(* Logix 5000 project; controller FV vendor 1 type 14 code 217 rev 31.11; software revision 31.00; part 54 of 63 *)
(* tags used below, declared in another part *)
   Alarm_Reset : BOOL;
   CWD : CHECKWORD_FLAGS;
   Default_Check_Time : DINT;
   Dummy : BOOL;
   FV_AV1 : PlantItem;   // AV1
   FV_AV1_ALARM : ALARM_DIGITAL;
   FV_AV1_C : ALIAS FOR Remote_IO:6:I.Data.4;   // YSV 1 outlet valve closed f/b
   FV_AV1_DR : ALIAS FOR Remote_IO:5:O.Data.0;   // YSV 1 outlet valve
   FV_AV1_O : ALIAS FOR Remote_IO:6:I.Data.0;   // YSV 1 outlet valve open f/b
   FV_AV1A : PlantItem;   // AV1A
   FV_AV1A_ALARM : ALARM_DIGITAL;
   FV_AV1A_C : ALIAS FOR Remote_IO:6:I.Data.10;   // AV1A seat clean valve closed f/b
   FV_AV1A_DR : ALIAS FOR Remote_IO:5:O.Data.4;   // AV1 seat clean valve
   FV_AV1A_O : ALIAS FOR Remote_IO:6:I.Data.8;   // AV1A seat clean valve open f/b
   FV_AV2 : PlantItem;   // AV2
   FV_AV2_ALARM : ALARM_DIGITAL;
   FV_AV2_C : ALIAS FOR Remote_IO:6:I.Data.5;   // Water flush valve closed f/b
   FV_AV2_DR : ALIAS FOR Remote_IO:5:O.Data.1;   // Water flush valve
   FV_AV2_O : ALIAS FOR Remote_IO:6:I.Data.1;   // Water flush valve open f/b
   FV_AV3 : PlantItem;   // AV3
   FV_AV3_ALARM : ALARM_DIGITAL;
   FV_AV3_C : ALIAS FOR Remote_IO:6:I.Data.6;   // CIP delivery valve closed f/b
   FV_AV3_DR : ALIAS FOR Remote_IO:5:O.Data.2;   // CIP delivery valve
   FV_AV3_O : ALIAS FOR Remote_IO:6:I.Data.2;   // CIP delivery valve open f/b
   FV_AV4 : PlantItem;   // AV4
   FV_AV4_ALARM : ALARM_DIGITAL;
   FV_AV4_C : ALIAS FOR Remote_IO:6:I.Data.7;   // Centrifuge main closed f/b
   FV_AV4_DR : ALIAS FOR Remote_IO:5:O.Data.3;   // Centrifuge main valve
   FV_AV4_O : ALIAS FOR Remote_IO:6:I.Data.3;   // Centrifuge main valve f/b
   FV_AV4A : PlantItem;   // AV4A
   FV_AV4A_ALARM : ALARM_DIGITAL;
   FV_AV4A_C : ALIAS FOR Remote_IO:6:I.Data.11;   // AV4A seat clean valve closed f/b
   FV_AV4A_DR : ALIAS FOR Remote_IO:5:O.Data.5;   // AV4 seat clean valve
   FV_AV4A_O : ALIAS FOR Remote_IO:6:I.Data.9;   // AV4A seat clean valve closed f/b
   FV_AV5 : PlantItem;   // AV5
   FV_AV5_ALARM : ALARM_DIGITAL;
   FV_AV5_C : ALIAS FOR Remote_IO:7:I.Data.9;
   FV_AV5_DR : ALIAS FOR Remote_IO:9:O.Data.12;
   FV_AV5_O : ALIAS FOR Remote_IO:7:I.Data.8;
   FV_B17 : INT[255];   // VES_ACTIVE Vessel active flags
   fv_bit_data_file_address : INT;
   fv_bit_file_bit_offset : INT;
   fv_bit_file_word_offset : INT;
   fv_bit_offset : INT;
   fv_bit_value_to_set : INT;
   FV_data_file_address : INT;
   FV_N110 : INT[255];   // FV DATA 0 CURRENT FV DATA
   FV_N111 : INT[50];   // FV1, CURRENT FV DATA
   FV_N112 : INT[50];   // FV2, CURRENT FV DATA
   FV_N113 : INT[50];   // FV3, CURRENT FV DATA
   FV_N114 : INT[50];   // FV4, CURRENT FV DATA
   FV_N115 : INT[50];   // FV5, CURRENT FV DATA
   FV_N116 : INT[50];   // FV6, CURRENT FV DATA
   FV_N117 : INT[50];   // FV7, CURRENT FV DATA
   FV_N118 : INT[50];   // FV8, CURRENT FV DATA
   FV_N119 : INT[50];   // FV9, CURRENT FV DATA
   FV_N120 : INT[50];   // FV10, CURRENT FV DATA
   FV_N121 : INT[50];   // FV11, CURRENT FV DATA
   FV_N122 : INT[50];   // FV12, CURRENT FV DATA
   FV_N123 : INT[50];   // FV13, CURRENT FV DATA
   FV_N124 : INT[50];   // FV14, CURRENT FV DATA
   FV_N125 : INT[50];   // FV15, CURRENT FV DATA
   FV_N126 : INT[50];   // FV16, CURRENT FV DATA
   FV_N127 : INT[50];   // FV17, CURRENT FV DATA
   FV_N128 : INT[50];   // FV18, CURRENT FV DATA
   FV_N129 : INT[50];   // FV19, CURRENT FV DATA
   FV_N130 : INT[50];   // FV20, CURRENT FV DATA
   FV_N131 : INT[50];   // FV21, CURRENT FV DATA
   FV_N132 : INT[50];   // FV22, CURRENT FV DATA
   FV_N133 : INT[50];   // FV23, CURRENT FV DATA
   FV_N134 : INT[50];   // FV24, CURRENT FV DATA
   FV_N135 : INT[50];   // FV25, CURRENT FV DATA
   FV_N136 : INT[50];   // YSV1, CURRENT FV DATA
   FV_N137 : INT[50];   // YSV2, CURRENT FV DATA
   FV_N138 : INT[50];   // YSV3, CURRENT FV DATA
   FV_N139 : INT[255];   // YST1
   FV_N140 : INT[255];   // YST2
   FV_N141 : INT[255];   // YSV1 DATA
   FV_N142 : INT[255];   // YSV2 DATA
   FV_N143 : INT[255];   // YSV3 DATA
   FV_N144 : INT[255];   // YST1 DATA
   FV_N145 : INT[255];   // YST2 DATA
   FV_N146 : INT[50];   // FV26, CURRENT FV DATA
   FV_N147 : INT[50];   // FV27, CURRENT FV DATA
   FV_N148 : INT[50];   // FV28, CURRENT FV DATA
   FV_N149 : INT[50];   // FV29, CURRENT FV DATA
   FV_N150 : INT[50];   // FV30, CURRENT FV DATA
   FV_N151 : INT[50];   // FV31, CURRENT FV DATA
   FV_R2V1 : PlantItem;   // R2V1
   FV_R2V1_ALARM : ALARM_DIGITAL;
   FV_R2V1_C : ALIAS FOR Remote_IO:7:I.Data.6;
   FV_R2V1_DR : ALIAS FOR Remote_IO:5:O.Data.10;
   FV_R2V1_O : ALIAS FOR Remote_IO:7:I.Data.2;
   FV_R2V2 : PlantItem;   // R2V2
   FV_R2V2_ALARM : ALARM_DIGITAL;
   FV_R2V2_C : ALIAS FOR Remote_IO:7:I.Data.7;
   FV_R2V2_DR : ALIAS FOR Remote_IO:5:O.Data.11;
   FV_R2V2_O : ALIAS FOR Remote_IO:7:I.Data.3;
   FV_value_to_set : INT;
   FV_word_offset : INT;
   FV_WYTR1 : PlantItem;   // WYTR1
   FV_WYTR1_ALARM : ALARM_DIGITAL;
   FV_WYTR1_C : ALIAS FOR Remote_IO:7:I.Data.4;
   FV_WYTR1_DR : ALIAS FOR Remote_IO:5:O.Data.8;
   FV_WYTR1_O : ALIAS FOR Remote_IO:7:I.Data.0;
   FV_WYTR2 : PlantItem;   // WYTR2
   FV_WYTR2_ALARM : ALARM_DIGITAL;
   FV_WYTR2_C : ALIAS FOR Remote_IO:7:I.Data.5;
   FV_WYTR2_DR : ALIAS FOR Remote_IO:5:O.Data.9;
   FV_WYTR2_O : ALIAS FOR Remote_IO:7:I.Data.1;
   Item_Faults_Are_Latched : BOOL;
   Item_Simulation_Flag : BOOL;
   One_Second_One_Scan : ALIAS FOR One_Second_1_scan;
   Scada_Valve_Fault_No : DINT;
   YP_AV2 : PlantItem;   // AV2
   YP_AV2_ALARM : ALARM_DIGITAL;
   YP_AV2_DR : ALIAS FOR RIO_Rack_3:3:O.Data.5;
   YP_AV2_O : ALIAS FOR RIO_Rack_3:1:I.Data.2;
(* FV_Common, continued *)

ROUTINE FV_Set_FV_Datafile_Value   (* ladder *)
   // Routine to Set the value of something within the FV Data Files, Used to replace indirection originally used
   0: SBR(FV_value_to_set,FV_data_file_address,FV_word_offset)OTE(Dummy);
   1: EQU(FV_data_file_address,110)MOV(FV_value_to_set,FV_N110[FV_word_offset]);
   2: EQU(FV_data_file_address,111)MOV(FV_value_to_set,FV_N111[FV_word_offset]);
   3: EQU(FV_data_file_address,112)MOV(FV_value_to_set,FV_N112[FV_word_offset]);
   4: EQU(FV_data_file_address,113)MOV(FV_value_to_set,FV_N113[FV_word_offset]);
   5: EQU(FV_data_file_address,114)MOV(FV_value_to_set,FV_N114[FV_word_offset]);
   6: EQU(FV_data_file_address,115)MOV(FV_value_to_set,FV_N115[FV_word_offset]);
   7: EQU(FV_data_file_address,116)MOV(FV_value_to_set,FV_N116[FV_word_offset]);
   8: EQU(FV_data_file_address,117)MOV(FV_value_to_set,FV_N117[FV_word_offset]);
   9: EQU(FV_data_file_address,118)MOV(FV_value_to_set,FV_N118[FV_word_offset]);
   10: EQU(FV_data_file_address,119)MOV(FV_value_to_set,FV_N119[FV_word_offset]);
   11: EQU(FV_data_file_address,120)MOV(FV_value_to_set,FV_N120[FV_word_offset]);
   12: EQU(FV_data_file_address,121)MOV(FV_value_to_set,FV_N121[FV_word_offset]);
   13: EQU(FV_data_file_address,122)MOV(FV_value_to_set,FV_N122[FV_word_offset]);
   14: EQU(FV_data_file_address,123)MOV(FV_value_to_set,FV_N123[FV_word_offset]);
   15: EQU(FV_data_file_address,124)MOV(FV_value_to_set,FV_N124[FV_word_offset]);
   16: EQU(FV_data_file_address,125)MOV(FV_value_to_set,FV_N125[FV_word_offset]);
   17: EQU(FV_data_file_address,126)MOV(FV_value_to_set,FV_N126[FV_word_offset]);
   18: EQU(FV_data_file_address,127)MOV(FV_value_to_set,FV_N127[FV_word_offset]);
   19: EQU(FV_data_file_address,128)MOV(FV_value_to_set,FV_N128[FV_word_offset]);
   20: EQU(FV_data_file_address,129)MOV(FV_value_to_set,FV_N129[FV_word_offset]);
   21: EQU(FV_data_file_address,130)MOV(FV_value_to_set,FV_N130[FV_word_offset]);
   22: EQU(FV_data_file_address,131)MOV(FV_value_to_set,FV_N131[FV_word_offset]);
   23: EQU(FV_data_file_address,132)MOV(FV_value_to_set,FV_N132[FV_word_offset]);
   24: EQU(FV_data_file_address,133)MOV(FV_value_to_set,FV_N133[FV_word_offset]);
   25: EQU(FV_data_file_address,134)MOV(FV_value_to_set,FV_N134[FV_word_offset]);
   26: EQU(FV_data_file_address,135)MOV(FV_value_to_set,FV_N135[FV_word_offset]);
   27: EQU(FV_data_file_address,136)MOV(FV_value_to_set,FV_N136[FV_word_offset]);
   28: EQU(FV_data_file_address,137)MOV(FV_value_to_set,FV_N137[FV_word_offset]);
   29: EQU(FV_data_file_address,138)MOV(FV_value_to_set,FV_N138[FV_word_offset]);
   30: EQU(FV_data_file_address,139)MOV(FV_value_to_set,FV_N139[FV_word_offset]);
   31: EQU(FV_data_file_address,140)MOV(FV_value_to_set,FV_N140[FV_word_offset]);
   32: EQU(FV_data_file_address,141)MOV(FV_value_to_set,FV_N141[FV_word_offset]);
   33: EQU(FV_data_file_address,142)MOV(FV_value_to_set,FV_N142[FV_word_offset]);
   34: EQU(FV_data_file_address,143)MOV(FV_value_to_set,FV_N143[FV_word_offset]);
   35: EQU(FV_data_file_address,144)MOV(FV_value_to_set,FV_N144[FV_word_offset]);
   36: EQU(FV_data_file_address,145)MOV(FV_value_to_set,FV_N145[FV_word_offset]);
   37: EQU(FV_data_file_address,146)MOV(FV_value_to_set,FV_N146[FV_word_offset]);
   38: EQU(FV_data_file_address,147)MOV(FV_value_to_set,FV_N147[FV_word_offset]);
   39: EQU(FV_data_file_address,148)MOV(FV_value_to_set,FV_N148[FV_word_offset]);
   40: EQU(FV_data_file_address,149)MOV(FV_value_to_set,FV_N149[FV_word_offset]);
   41: EQU(FV_data_file_address,150)MOV(FV_value_to_set,FV_N150[FV_word_offset]);
   42: EQU(FV_data_file_address,151)MOV(FV_value_to_set,FV_N151[FV_word_offset]);
   43: RET();
END_ROUTINE

ROUTINE FV_SetBitFile_Value   (* ladder *)
   // Sets the Value of a bit within a bit file, Can use complete bit offset across words
   0: SBR(fv_bit_value_to_set,fv_bit_data_file_address,fv_bit_offset)OTE(Dummy);
   1: DIV(fv_bit_offset,16,fv_bit_file_word_offset)MOD(fv_bit_offset,16,fv_bit_file_bit_offset);
   // Bit File 17
   2: EQU(fv_bit_data_file_address,17)[EQU(fv_bit_value_to_set,1) OTL(FV_B17[fv_bit_file_word_offset].[fv_bit_file_bit_offset]) ,EQU(fv_bit_value_to_set,0) OTU(FV_B17[fv_bit_file_word_offset].[fv_bit_file_bit_offset]) ];
   3: RET();
END_ROUTINE

ROUTINE FV_Valves   (* ladder *)
   0: [NEQ(FV_AV1.DriveBits,0) OTE(FV_AV1.CW.[CWD.AUTODRV]) ,[XIC(FV_AV1.CW.[CWD.AUTODRV]) XIO(FV_AV1.CW.[CWD.MANUAL]) ,XIC(FV_AV1.CW.[CWD.MANDRV]) XIC(FV_AV1.CW.[CWD.MANUAL]) ] OTE(FV_AV1.CW.[CWD.OUTPUT]) ,XIC(FV_AV1.CW.[CWD.OUTPUT]) OTE(FV_AV1_DR) ,XIC(S:FS) [OTU(FV_AV1.CW.[CWD.MANUAL]) ,LEQ(FV_AV1.CheckTime,0) MOV(Default_Check_Time,FV_AV1.CheckTime) ] ,[[XIC(FV_AV1_O) XIO(Item_Simulation_Flag) ,XIC(Item_Simulation_Flag) XIC(FV_AV1.CW.[CWD.OUTPUT]) XIO(FV_AV1.CW.[CWD.SIMFAIL]) ] OTE(FV_AV1.CW.[CWD.OPENFB]) ,[XIC(FV_AV1_C) XIO(Item_Simulation_Flag) ,XIC(Item_Simulation_Flag) XIO(FV_AV1.CW.[CWD.OUTPUT]) XIO(FV_AV1.CW.[CWD.SIMFAIL]) ] OTE(FV_AV1.CW.[CWD.CLOSEDFB]) ] ,[XIC(FV_AV1.CW.[CWD.OUTPUT]) XIO(FV_AV1.CW.[CWD.PREVSCAN]) ,XIO(FV_AV1.CW.[CWD.OUTPUT]) XIC(FV_AV1.CW.[CWD.PREVSCAN]) ] CLR(FV_AV1.CheckTimer) ,XIC(One_Second_One_Scan) LES(FV_AV1.CheckTimer,FV_AV1.CheckTime) ADD(FV_AV1.CheckTimer,1,FV_AV1.CheckTimer) ,XIO(FV_AV1.CW.[CWD.FAULT]) OTU(FV_AV1.CW.[CWD.FAULTLOGGED]) ,[GEQ(FV_AV1.CheckTimer,FV_AV1.CheckTime) [XIC(FV_AV1.CW.[CWD.OUTPUT]) [XIO(FV_AV1.CW.[CWD.OPENFB]) ,XIC(FV_AV1.CW.[CWD.CLOSEDFB]) ] ,XIO(FV_AV1.CW.[CWD.OUTPUT]) [XIC(FV_AV1.CW.[CWD.OPENFB]) ,XIO(FV_AV1.CW.[CWD.CLOSEDFB]) ] ] ,XIC(FV_AV1.CW.[CWD.FAULT]) XIC(Item_Faults_Are_Latched) ,XIC(FV_AV1.CW.[CWD.HIGHLIGHT]) ] XIO(FV_AV1.CW.[CWD.CHECKOFF]) XIO(Alarm_Reset) [OTE(FV_AV1.CW.[CWD.FAULT]) ,ALMD(FV_AV1_ALARM,0,0,0,0) ] ,XIC(FV_AV1.CW.[CWD.OUTPUT]) OTE(FV_AV1.CW.[CWD.PREVSCAN]) ,XIC(FV_AV1.CW.[CWD.FAULT]) EQU(Scada_Valve_Fault_No,0) XIO(FV_AV1.CW.[CWD.FAULTLOGGED]) [MOV(10001,Scada_Valve_Fault_No) ,OTL(FV_AV1.CW.[CWD.FAULTLOGGED]) ] ];
   1: [NEQ(FV_AV2.DriveBits,0) OTE(FV_AV2.CW.[CWD.AUTODRV]) ,[XIC(FV_AV2.CW.[CWD.AUTODRV]) XIO(FV_AV2.CW.[CWD.MANUAL]) ,XIC(FV_AV2.CW.[CWD.MANDRV]) XIC(FV_AV2.CW.[CWD.MANUAL]) ] OTE(FV_AV2.CW.[CWD.OUTPUT]) ,XIC(FV_AV2.CW.[CWD.OUTPUT]) OTE(FV_AV2_DR) ,XIC(S:FS) [OTU(FV_AV2.CW.[CWD.MANUAL]) ,LEQ(FV_AV2.CheckTime,0) MOV(Default_Check_Time,FV_AV2.CheckTime) ] ,[[XIC(FV_AV2_O) XIO(Item_Simulation_Flag) ,XIC(Item_Simulation_Flag) XIC(FV_AV2.CW.[CWD.OUTPUT]) XIO(FV_AV2.CW.[CWD.SIMFAIL]) ] OTE(FV_AV2.CW.[CWD.OPENFB]) ,[XIC(FV_AV2_C) XIO(Item_Simulation_Flag) ,XIC(Item_Simulation_Flag) XIO(FV_AV2.CW.[CWD.OUTPUT]) XIO(FV_AV2.CW.[CWD.SIMFAIL]) ] OTE(FV_AV2.CW.[CWD.CLOSEDFB]) ] ,[XIC(FV_AV2.CW.[CWD.OUTPUT]) XIO(FV_AV2.CW.[CWD.PREVSCAN]) ,XIO(FV_AV2.CW.[CWD.OUTPUT]) XIC(FV_AV2.CW.[CWD.PREVSCAN]) ] CLR(FV_AV2.CheckTimer) ,XIC(One_Second_One_Scan) LES(FV_AV2.CheckTimer,FV_AV2.CheckTime) ADD(FV_AV2.CheckTimer,1,FV_AV2.CheckTimer) ,XIO(FV_AV2.CW.[CWD.FAULT]) OTU(FV_AV2.CW.[CWD.FAULTLOGGED]) ,[GEQ(FV_AV2.CheckTimer,FV_AV2.CheckTime) [XIC(FV_AV2.CW.[CWD.OUTPUT]) [XIO(FV_AV2.CW.[CWD.OPENFB]) ,XIC(FV_AV2.CW.[CWD.CLOSEDFB]) ] ,XIO(FV_AV2.CW.[CWD.OUTPUT]) [XIC(FV_AV2.CW.[CWD.OPENFB]) ,XIO(FV_AV2.CW.[CWD.CLOSEDFB]) ] ] ,XIC(FV_AV2.CW.[CWD.FAULT]) XIC(Item_Faults_Are_Latched) ,XIC(FV_AV2.CW.[CWD.HIGHLIGHT]) ] XIO(FV_AV2.CW.[CWD.CHECKOFF]) XIO(Alarm_Reset) [OTE(FV_AV2.CW.[CWD.FAULT]) ,ALMD(FV_AV2_ALARM,0,0,0,0) ] ,XIC(FV_AV2.CW.[CWD.OUTPUT]) OTE(FV_AV2.CW.[CWD.PREVSCAN]) ,XIC(FV_AV2.CW.[CWD.FAULT]) EQU(Scada_Valve_Fault_No,0) XIO(FV_AV2.CW.[CWD.FAULTLOGGED]) [MOV(10001,Scada_Valve_Fault_No) ,OTL(FV_AV2.CW.[CWD.FAULTLOGGED]) ] ];
   2: [NEQ(FV_AV3.DriveBits,0) OTE(FV_AV3.CW.[CWD.AUTODRV]) ,[XIC(FV_AV3.CW.[CWD.AUTODRV]) XIO(FV_AV3.CW.[CWD.MANUAL]) ,XIC(FV_AV3.CW.[CWD.MANDRV]) XIC(FV_AV3.CW.[CWD.MANUAL]) ] OTE(FV_AV3.CW.[CWD.OUTPUT]) ,XIC(FV_AV3.CW.[CWD.OUTPUT]) OTE(FV_AV3_DR) ,XIC(S:FS) [OTU(FV_AV3.CW.[CWD.MANUAL]) ,LEQ(FV_AV3.CheckTime,0) MOV(Default_Check_Time,FV_AV3.CheckTime) ] ,[[XIC(FV_AV3_O) XIO(Item_Simulation_Flag) ,XIC(Item_Simulation_Flag) XIC(FV_AV3.CW.[CWD.OUTPUT]) XIO(FV_AV3.CW.[CWD.SIMFAIL]) ] OTE(FV_AV3.CW.[CWD.OPENFB]) ,[XIC(FV_AV3_C) XIO(Item_Simulation_Flag) ,XIC(Item_Simulation_Flag) XIO(FV_AV3.CW.[CWD.OUTPUT]) XIO(FV_AV3.CW.[CWD.SIMFAIL]) ] OTE(FV_AV3.CW.[CWD.CLOSEDFB]) ] ,[XIC(FV_AV3.CW.[CWD.OUTPUT]) XIO(FV_AV3.CW.[CWD.PREVSCAN]) ,XIO(FV_AV3.CW.[CWD.OUTPUT]) XIC(FV_AV3.CW.[CWD.PREVSCAN]) ] CLR(FV_AV3.CheckTimer) ,XIC(One_Second_One_Scan) LES(FV_AV3.CheckTimer,FV_AV3.CheckTime) ADD(FV_AV3.CheckTimer,1,FV_AV3.CheckTimer) ,XIO(FV_AV3.CW.[CWD.FAULT]) OTU(FV_AV3.CW.[CWD.FAULTLOGGED]) ,[GEQ(FV_AV3.CheckTimer,FV_AV3.CheckTime) [XIC(FV_AV3.CW.[CWD.OUTPUT]) [XIO(FV_AV3.CW.[CWD.OPENFB]) ,XIC(FV_AV3.CW.[CWD.CLOSEDFB]) ] ,XIO(FV_AV3.CW.[CWD.OUTPUT]) [XIC(FV_AV3.CW.[CWD.OPENFB]) ,XIO(FV_AV3.CW.[CWD.CLOSEDFB]) ] ] ,XIC(FV_AV3.CW.[CWD.FAULT]) XIC(Item_Faults_Are_Latched) ,XIC(FV_AV3.CW.[CWD.HIGHLIGHT]) ] XIO(FV_AV3.CW.[CWD.CHECKOFF]) XIO(Alarm_Reset) [OTE(FV_AV3.CW.[CWD.FAULT]) ,ALMD(FV_AV3_ALARM,0,0,0,0) ] ,XIC(FV_AV3.CW.[CWD.OUTPUT]) OTE(FV_AV3.CW.[CWD.PREVSCAN]) ,XIC(FV_AV3.CW.[CWD.FAULT]) EQU(Scada_Valve_Fault_No,0) XIO(FV_AV3.CW.[CWD.FAULTLOGGED]) [MOV(10001,Scada_Valve_Fault_No) ,OTL(FV_AV3.CW.[CWD.FAULTLOGGED]) ] ];
   3: [NEQ(FV_AV4.DriveBits,0) OTE(FV_AV4.CW.[CWD.AUTODRV]) ,[XIC(FV_AV4.CW.[CWD.AUTODRV]) XIO(FV_AV4.CW.[CWD.MANUAL]) ,XIC(FV_AV4.CW.[CWD.MANDRV]) XIC(FV_AV4.CW.[CWD.MANUAL]) ] OTE(FV_AV4.CW.[CWD.OUTPUT]) ,XIC(FV_AV4.CW.[CWD.OUTPUT]) OTE(FV_AV4_DR) ,XIC(S:FS) [OTU(FV_AV4.CW.[CWD.MANUAL]) ,LEQ(FV_AV4.CheckTime,0) MOV(Default_Check_Time,FV_AV4.CheckTime) ] ,[[XIC(FV_AV4_O) XIO(Item_Simulation_Flag) ,XIC(Item_Simulation_Flag) XIC(FV_AV4.CW.[CWD.OUTPUT]) XIO(FV_AV4.CW.[CWD.SIMFAIL]) ] OTE(FV_AV4.CW.[CWD.OPENFB]) ,[XIC(FV_AV4_C) XIO(Item_Simulation_Flag) ,XIC(Item_Simulation_Flag) XIO(FV_AV4.CW.[CWD.OUTPUT]) XIO(FV_AV4.CW.[CWD.SIMFAIL]) ] OTE(FV_AV4.CW.[CWD.CLOSEDFB]) ] ,[XIC(FV_AV4.CW.[CWD.OUTPUT]) XIO(FV_AV4.CW.[CWD.PREVSCAN]) ,XIO(FV_AV4.CW.[CWD.OUTPUT]) XIC(FV_AV4.CW.[CWD.PREVSCAN]) ] CLR(FV_AV4.CheckTimer) ,XIC(One_Second_One_Scan) LES(FV_AV4.CheckTimer,FV_AV4.CheckTime) ADD(FV_AV4.CheckTimer,1,FV_AV4.CheckTimer) ,XIO(FV_AV4.CW.[CWD.FAULT]) OTU(FV_AV4.CW.[CWD.FAULTLOGGED]) ,[GEQ(FV_AV4.CheckTimer,FV_AV4.CheckTime) [XIC(FV_AV4.CW.[CWD.OUTPUT]) [XIO(FV_AV4.CW.[CWD.OPENFB]) ,XIC(FV_AV4.CW.[CWD.CLOSEDFB]) ] ,XIO(FV_AV4.CW.[CWD.OUTPUT]) [XIC(FV_AV4.CW.[CWD.OPENFB]) ,XIO(FV_AV4.CW.[CWD.CLOSEDFB]) ] ] ,XIC(FV_AV4.CW.[CWD.FAULT]) XIC(Item_Faults_Are_Latched) ,XIC(FV_AV4.CW.[CWD.HIGHLIGHT]) ] XIO(FV_AV4.CW.[CWD.CHECKOFF]) XIO(Alarm_Reset) [OTE(FV_AV4.CW.[CWD.FAULT]) ,ALMD(FV_AV4_ALARM,0,0,0,0) ] ,XIC(FV_AV4.CW.[CWD.OUTPUT]) OTE(FV_AV4.CW.[CWD.PREVSCAN]) ,XIC(FV_AV4.CW.[CWD.FAULT]) EQU(Scada_Valve_Fault_No,0) XIO(FV_AV4.CW.[CWD.FAULTLOGGED]) [MOV(10001,Scada_Valve_Fault_No) ,OTL(FV_AV4.CW.[CWD.FAULTLOGGED]) ] ];
   4: [NEQ(FV_AV1A.DriveBits,0) OTE(FV_AV1A.CW.[CWD.AUTODRV]) ,[XIC(FV_AV1A.CW.[CWD.AUTODRV]) XIO(FV_AV1A.CW.[CWD.MANUAL]) ,XIC(FV_AV1A.CW.[CWD.MANDRV]) XIC(FV_AV1A.CW.[CWD.MANUAL]) ] OTE(FV_AV1A.CW.[CWD.OUTPUT]) ,XIC(FV_AV1A.CW.[CWD.OUTPUT]) OTE(FV_AV1A_DR) ,XIC(S:FS) [OTU(FV_AV1A.CW.[CWD.MANUAL]) ,LEQ(FV_AV1A.CheckTime,0) MOV(Default_Check_Time,FV_AV1A.CheckTime) ] ,[[XIC(FV_AV1A_O) XIO(Item_Simulation_Flag) ,XIC(Item_Simulation_Flag) XIC(FV_AV1A.CW.[CWD.OUTPUT]) XIO(FV_AV1A.CW.[CWD.SIMFAIL]) ] OTE(FV_AV1A.CW.[CWD.OPENFB]) ,[XIC(FV_AV1A_C) XIO(Item_Simulation_Flag) ,XIC(Item_Simulation_Flag) XIO(FV_AV1A.CW.[CWD.OUTPUT]) XIO(FV_AV1A.CW.[CWD.SIMFAIL]) ] OTE(FV_AV1A.CW.[CWD.CLOSEDFB]) ] ,[XIC(FV_AV1A.CW.[CWD.OUTPUT]) XIO(FV_AV1A.CW.[CWD.PREVSCAN]) ,XIO(FV_AV1A.CW.[CWD.OUTPUT]) XIC(FV_AV1A.CW.[CWD.PREVSCAN]) ] CLR(FV_AV1A.CheckTimer) ,XIC(One_Second_One_Scan) LES(FV_AV1A.CheckTimer,FV_AV1A.CheckTime) ADD(FV_AV1A.CheckTimer,1,FV_AV1A.CheckTimer) ,XIO(FV_AV1A.CW.[CWD.FAULT]) OTU(FV_AV1A.CW.[CWD.FAULTLOGGED]) ,[GEQ(FV_AV1A.CheckTimer,FV_AV1A.CheckTime) [XIC(FV_AV1A.CW.[CWD.OUTPUT]) [XIO(FV_AV1A.CW.[CWD.OPENFB]) ,XIC(FV_AV1A.CW.[CWD.CLOSEDFB]) ] ,XIO(FV_AV1A.CW.[CWD.OUTPUT]) [XIC(FV_AV1A.CW.[CWD.OPENFB]) ,XIO(FV_AV1A.CW.[CWD.CLOSEDFB]) ] ] ,XIC(FV_AV1A.CW.[CWD.FAULT]) XIC(Item_Faults_Are_Latched) ,XIC(FV_AV1A.CW.[CWD.HIGHLIGHT]) ] XIO(FV_AV1A.CW.[CWD.CHECKOFF]) XIO(Alarm_Reset) [OTE(FV_AV1A.CW.[CWD.FAULT]) ,ALMD(FV_AV1A_ALARM,0,0,0,0) ] ,XIC(FV_AV1A.CW.[CWD.OUTPUT]) OTE(FV_AV1A.CW.[CWD.PREVSCAN]) ,XIC(FV_AV1A.CW.[CWD.FAULT]) EQU(Scada_Valve_Fault_No,0) XIO(FV_AV1A.CW.[CWD.FAULTLOGGED]) [MOV(10001,Scada_Valve_Fault_No) ,OTL(FV_AV1A.CW.[CWD.FAULTLOGGED]) ] ];
   5: [NEQ(FV_AV4A.DriveBits,0) OTE(FV_AV4A.CW.[CWD.AUTODRV]) ,[XIC(FV_AV4A.CW.[CWD.AUTODRV]) XIO(FV_AV4A.CW.[CWD.MANUAL]) ,XIC(FV_AV4A.CW.[CWD.MANDRV]) XIC(FV_AV4A.CW.[CWD.MANUAL]) ] OTE(FV_AV4A.CW.[CWD.OUTPUT]) ,XIC(FV_AV4A.CW.[CWD.OUTPUT]) OTE(FV_AV4A_DR) ,XIC(S:FS) [OTU(FV_AV4A.CW.[CWD.MANUAL]) ,LEQ(FV_AV4A.CheckTime,0) MOV(Default_Check_Time,FV_AV4A.CheckTime) ] ,[[XIC(FV_AV4A_O) XIO(Item_Simulation_Flag) ,XIC(Item_Simulation_Flag) XIC(FV_AV4A.CW.[CWD.OUTPUT]) XIO(FV_AV4A.CW.[CWD.SIMFAIL]) ] OTE(FV_AV4A.CW.[CWD.OPENFB]) ,[XIC(FV_AV4A_C) XIO(Item_Simulation_Flag) ,XIC(Item_Simulation_Flag) XIO(FV_AV4A.CW.[CWD.OUTPUT]) XIO(FV_AV4A.CW.[CWD.SIMFAIL]) ] OTE(FV_AV4A.CW.[CWD.CLOSEDFB]) ] ,[XIC(FV_AV4A.CW.[CWD.OUTPUT]) XIO(FV_AV4A.CW.[CWD.PREVSCAN]) ,XIO(FV_AV4A.CW.[CWD.OUTPUT]) XIC(FV_AV4A.CW.[CWD.PREVSCAN]) ] CLR(FV_AV4A.CheckTimer) ,XIC(One_Second_One_Scan) LES(FV_AV4A.CheckTimer,FV_AV4A.CheckTime) ADD(FV_AV4A.CheckTimer,1,FV_AV4A.CheckTimer) ,XIO(FV_AV4A.CW.[CWD.FAULT]) OTU(FV_AV4A.CW.[CWD.FAULTLOGGED]) ,[GEQ(FV_AV4A.CheckTimer,FV_AV4A.CheckTime) [XIC(FV_AV4A.CW.[CWD.OUTPUT]) [XIO(FV_AV4A.CW.[CWD.OPENFB]) ,XIC(FV_AV4A.CW.[CWD.CLOSEDFB]) ] ,XIO(FV_AV4A.CW.[CWD.OUTPUT]) [XIC(FV_AV4A.CW.[CWD.OPENFB]) ,XIO(FV_AV4A.CW.[CWD.CLOSEDFB]) ] ] ,XIC(FV_AV4A.CW.[CWD.FAULT]) XIC(Item_Faults_Are_Latched) ,XIC(FV_AV4A.CW.[CWD.HIGHLIGHT]) ] XIO(FV_AV4A.CW.[CWD.CHECKOFF]) XIO(Alarm_Reset) [OTE(FV_AV4A.CW.[CWD.FAULT]) ,ALMD(FV_AV4A_ALARM,0,0,0,0) ] ,XIC(FV_AV4A.CW.[CWD.OUTPUT]) OTE(FV_AV4A.CW.[CWD.PREVSCAN]) ,XIC(FV_AV4A.CW.[CWD.FAULT]) EQU(Scada_Valve_Fault_No,0) XIO(FV_AV4A.CW.[CWD.FAULTLOGGED]) [MOV(10001,Scada_Valve_Fault_No) ,OTL(FV_AV4A.CW.[CWD.FAULTLOGGED]) ] ];
   6: [NEQ(FV_WYTR1.DriveBits,0) OTE(FV_WYTR1.CW.[CWD.AUTODRV]) ,[XIC(FV_WYTR1.CW.[CWD.AUTODRV]) XIO(FV_WYTR1.CW.[CWD.MANUAL]) ,XIC(FV_WYTR1.CW.[CWD.MANDRV]) XIC(FV_WYTR1.CW.[CWD.MANUAL]) ] OTE(FV_WYTR1.CW.[CWD.OUTPUT]) ,XIC(FV_WYTR1.CW.[CWD.OUTPUT]) OTE(FV_WYTR1_DR) ,XIC(S:FS) [OTU(FV_WYTR1.CW.[CWD.MANUAL]) ,LEQ(FV_WYTR1.CheckTime,0) MOV(Default_Check_Time,FV_WYTR1.CheckTime) ] ,[[XIC(FV_WYTR1_O) XIO(Item_Simulation_Flag) ,XIC(Item_Simulation_Flag) XIC(FV_WYTR1.CW.[CWD.OUTPUT]) XIO(FV_WYTR1.CW.[CWD.SIMFAIL]) ] OTE(FV_WYTR1.CW.[CWD.OPENFB]) ,[XIC(FV_WYTR1_C) XIO(Item_Simulation_Flag) ,XIC(Item_Simulation_Flag) XIO(FV_WYTR1.CW.[CWD.OUTPUT]) XIO(FV_WYTR1.CW.[CWD.SIMFAIL]) ] OTE(FV_WYTR1.CW.[CWD.CLOSEDFB]) ] ,[XIC(FV_WYTR1.CW.[CWD.OUTPUT]) XIO(FV_WYTR1.CW.[CWD.PREVSCAN]) ,XIO(FV_WYTR1.CW.[CWD.OUTPUT]) XIC(FV_WYTR1.CW.[CWD.PREVSCAN]) ] CLR(FV_WYTR1.CheckTimer) ,XIC(One_Second_One_Scan) LES(FV_WYTR1.CheckTimer,FV_WYTR1.CheckTime) ADD(FV_WYTR1.CheckTimer,1,FV_WYTR1.CheckTimer) ,XIO(FV_WYTR1.CW.[CWD.FAULT]) OTU(FV_WYTR1.CW.[CWD.FAULTLOGGED]) ,[GEQ(FV_WYTR1.CheckTimer,FV_WYTR1.CheckTime) [XIC(FV_WYTR1.CW.[CWD.OUTPUT]) [XIO(FV_WYTR1.CW.[CWD.OPENFB]) ,XIC(FV_WYTR1.CW.[CWD.CLOSEDFB]) ] ,XIO(FV_WYTR1.CW.[CWD.OUTPUT]) [XIC(FV_WYTR1.CW.[CWD.OPENFB]) ,XIO(FV_WYTR1.CW.[CWD.CLOSEDFB]) ] ] ,XIC(FV_WYTR1.CW.[CWD.FAULT]) XIC(Item_Faults_Are_Latched) ,XIC(FV_WYTR1.CW.[CWD.HIGHLIGHT]) ] XIO(FV_WYTR1.CW.[CWD.CHECKOFF]) XIO(Alarm_Reset) [OTE(FV_WYTR1.CW.[CWD.FAULT]) ,ALMD(FV_WYTR1_ALARM,0,0,0,0) ] ,XIC(FV_WYTR1.CW.[CWD.OUTPUT]) OTE(FV_WYTR1.CW.[CWD.PREVSCAN]) ,XIC(FV_WYTR1.CW.[CWD.FAULT]) EQU(Scada_Valve_Fault_No,0) XIO(FV_WYTR1.CW.[CWD.FAULTLOGGED]) [MOV(10001,Scada_Valve_Fault_No) ,OTL(FV_WYTR1.CW.[CWD.FAULTLOGGED]) ] ];
   7: [NEQ(FV_WYTR2.DriveBits,0) OTE(FV_WYTR2.CW.[CWD.AUTODRV]) ,[XIC(FV_WYTR2.CW.[CWD.AUTODRV]) XIO(FV_WYTR2.CW.[CWD.MANUAL]) ,XIC(FV_WYTR2.CW.[CWD.MANDRV]) XIC(FV_WYTR2.CW.[CWD.MANUAL]) ] OTE(FV_WYTR2.CW.[CWD.OUTPUT]) ,XIC(FV_WYTR2.CW.[CWD.OUTPUT]) OTE(FV_WYTR2_DR) ,XIC(S:FS) [OTU(FV_WYTR2.CW.[CWD.MANUAL]) ,LEQ(FV_WYTR2.CheckTime,0) MOV(Default_Check_Time,FV_WYTR2.CheckTime) ] ,[[XIC(FV_WYTR2_O) XIO(Item_Simulation_Flag) ,XIC(Item_Simulation_Flag) XIC(FV_WYTR2.CW.[CWD.OUTPUT]) XIO(FV_WYTR2.CW.[CWD.SIMFAIL]) ] OTE(FV_WYTR2.CW.[CWD.OPENFB]) ,[XIC(FV_WYTR2_C) XIO(Item_Simulation_Flag) ,XIC(Item_Simulation_Flag) XIO(FV_WYTR2.CW.[CWD.OUTPUT]) XIO(FV_WYTR2.CW.[CWD.SIMFAIL]) ] OTE(FV_WYTR2.CW.[CWD.CLOSEDFB]) ] ,[XIC(FV_WYTR2.CW.[CWD.OUTPUT]) XIO(FV_WYTR2.CW.[CWD.PREVSCAN]) ,XIO(FV_WYTR2.CW.[CWD.OUTPUT]) XIC(FV_WYTR2.CW.[CWD.PREVSCAN]) ] CLR(FV_WYTR2.CheckTimer) ,XIC(One_Second_One_Scan) LES(FV_WYTR2.CheckTimer,FV_WYTR2.CheckTime) ADD(FV_WYTR2.CheckTimer,1,FV_WYTR2.CheckTimer) ,XIO(FV_WYTR2.CW.[CWD.FAULT]) OTU(FV_WYTR2.CW.[CWD.FAULTLOGGED]) ,[GEQ(FV_WYTR2.CheckTimer,FV_WYTR2.CheckTime) [XIC(FV_WYTR2.CW.[CWD.OUTPUT]) [XIO(FV_WYTR2.CW.[CWD.OPENFB]) ,XIC(FV_WYTR2.CW.[CWD.CLOSEDFB]) ] ,XIO(FV_WYTR2.CW.[CWD.OUTPUT]) [XIC(FV_WYTR2.CW.[CWD.OPENFB]) ,XIO(FV_WYTR2.CW.[CWD.CLOSEDFB]) ] ] ,XIC(FV_WYTR2.CW.[CWD.FAULT]) XIC(Item_Faults_Are_Latched) ,XIC(FV_WYTR2.CW.[CWD.HIGHLIGHT]) ] XIO(FV_WYTR2.CW.[CWD.CHECKOFF]) XIO(Alarm_Reset) [OTE(FV_WYTR2.CW.[CWD.FAULT]) ,ALMD(FV_WYTR2_ALARM,0,0,0,0) ] ,XIC(FV_WYTR2.CW.[CWD.OUTPUT]) OTE(FV_WYTR2.CW.[CWD.PREVSCAN]) ,XIC(FV_WYTR2.CW.[CWD.FAULT]) EQU(Scada_Valve_Fault_No,0) XIO(FV_WYTR2.CW.[CWD.FAULTLOGGED]) [MOV(10001,Scada_Valve_Fault_No) ,OTL(FV_WYTR2.CW.[CWD.FAULTLOGGED]) ] ];
   8: [NEQ(FV_R2V1.DriveBits,0) OTE(FV_R2V1.CW.[CWD.AUTODRV]) ,[XIC(FV_R2V1.CW.[CWD.AUTODRV]) XIO(FV_R2V1.CW.[CWD.MANUAL]) ,XIC(FV_R2V1.CW.[CWD.MANDRV]) XIC(FV_R2V1.CW.[CWD.MANUAL]) ] OTE(FV_R2V1.CW.[CWD.OUTPUT]) ,XIC(FV_R2V1.CW.[CWD.OUTPUT]) OTE(FV_R2V1_DR) ,XIC(S:FS) [OTU(FV_R2V1.CW.[CWD.MANUAL]) ,LEQ(FV_R2V1.CheckTime,0) MOV(Default_Check_Time,FV_R2V1.CheckTime) ] ,[[XIC(FV_R2V1_O) XIO(Item_Simulation_Flag) ,XIC(Item_Simulation_Flag) XIC(FV_R2V1.CW.[CWD.OUTPUT]) XIO(FV_R2V1.CW.[CWD.SIMFAIL]) ] OTE(FV_R2V1.CW.[CWD.OPENFB]) ,[XIC(FV_R2V1_C) XIO(Item_Simulation_Flag) ,XIC(Item_Simulation_Flag) XIO(FV_R2V1.CW.[CWD.OUTPUT]) XIO(FV_R2V1.CW.[CWD.SIMFAIL]) ] OTE(FV_R2V1.CW.[CWD.CLOSEDFB]) ] ,[XIC(FV_R2V1.CW.[CWD.OUTPUT]) XIO(FV_R2V1.CW.[CWD.PREVSCAN]) ,XIO(FV_R2V1.CW.[CWD.OUTPUT]) XIC(FV_R2V1.CW.[CWD.PREVSCAN]) ] CLR(FV_R2V1.CheckTimer) ,XIC(One_Second_One_Scan) LES(FV_R2V1.CheckTimer,FV_R2V1.CheckTime) ADD(FV_R2V1.CheckTimer,1,FV_R2V1.CheckTimer) ,XIO(FV_R2V1.CW.[CWD.FAULT]) OTU(FV_R2V1.CW.[CWD.FAULTLOGGED]) ,[GEQ(FV_R2V1.CheckTimer,FV_R2V1.CheckTime) [XIC(FV_R2V1.CW.[CWD.OUTPUT]) [XIO(FV_R2V1.CW.[CWD.OPENFB]) ,XIC(FV_R2V1.CW.[CWD.CLOSEDFB]) ] ,XIO(FV_R2V1.CW.[CWD.OUTPUT]) [XIC(FV_R2V1.CW.[CWD.OPENFB]) ,XIO(FV_R2V1.CW.[CWD.CLOSEDFB]) ] ] ,XIC(FV_R2V1.CW.[CWD.FAULT]) XIC(Item_Faults_Are_Latched) ,XIC(FV_R2V1.CW.[CWD.HIGHLIGHT]) ] XIO(FV_R2V1.CW.[CWD.CHECKOFF]) XIO(Alarm_Reset) [OTE(FV_R2V1.CW.[CWD.FAULT]) ,ALMD(FV_R2V1_ALARM,0,0,0,0) ] ,XIC(FV_R2V1.CW.[CWD.OUTPUT]) OTE(FV_R2V1.CW.[CWD.PREVSCAN]) ,XIC(FV_R2V1.CW.[CWD.FAULT]) EQU(Scada_Valve_Fault_No,0) XIO(FV_R2V1.CW.[CWD.FAULTLOGGED]) [MOV(10001,Scada_Valve_Fault_No) ,OTL(FV_R2V1.CW.[CWD.FAULTLOGGED]) ] ];
   9: [NEQ(FV_R2V2.DriveBits,0) OTE(FV_R2V2.CW.[CWD.AUTODRV]) ,[XIC(FV_R2V2.CW.[CWD.AUTODRV]) XIO(FV_R2V2.CW.[CWD.MANUAL]) ,XIC(FV_R2V2.CW.[CWD.MANDRV]) XIC(FV_R2V2.CW.[CWD.MANUAL]) ] OTE(FV_R2V2.CW.[CWD.OUTPUT]) ,XIC(FV_R2V2.CW.[CWD.OUTPUT]) OTE(FV_R2V2_DR) ,XIC(S:FS) [OTU(FV_R2V2.CW.[CWD.MANUAL]) ,LEQ(FV_R2V2.CheckTime,0) MOV(Default_Check_Time,FV_R2V2.CheckTime) ] ,[[XIC(FV_R2V2_O) XIO(Item_Simulation_Flag) ,XIC(Item_Simulation_Flag) XIC(FV_R2V2.CW.[CWD.OUTPUT]) XIO(FV_R2V2.CW.[CWD.SIMFAIL]) ] OTE(FV_R2V2.CW.[CWD.OPENFB]) ,[XIC(FV_R2V2_C) XIO(Item_Simulation_Flag) ,XIC(Item_Simulation_Flag) XIO(FV_R2V2.CW.[CWD.OUTPUT]) XIO(FV_R2V2.CW.[CWD.SIMFAIL]) ] OTE(FV_R2V2.CW.[CWD.CLOSEDFB]) ] ,[XIC(FV_R2V2.CW.[CWD.OUTPUT]) XIO(FV_R2V2.CW.[CWD.PREVSCAN]) ,XIO(FV_R2V2.CW.[CWD.OUTPUT]) XIC(FV_R2V2.CW.[CWD.PREVSCAN]) ] CLR(FV_R2V2.CheckTimer) ,XIC(One_Second_One_Scan) LES(FV_R2V2.CheckTimer,FV_R2V2.CheckTime) ADD(FV_R2V2.CheckTimer,1,FV_R2V2.CheckTimer) ,XIO(FV_R2V2.CW.[CWD.FAULT]) OTU(FV_R2V2.CW.[CWD.FAULTLOGGED]) ,[GEQ(FV_R2V2.CheckTimer,FV_R2V2.CheckTime) [XIC(FV_R2V2.CW.[CWD.OUTPUT]) [XIO(FV_R2V2.CW.[CWD.OPENFB]) ,XIC(FV_R2V2.CW.[CWD.CLOSEDFB]) ] ,XIO(FV_R2V2.CW.[CWD.OUTPUT]) [XIC(FV_R2V2.CW.[CWD.OPENFB]) ,XIO(FV_R2V2.CW.[CWD.CLOSEDFB]) ] ] ,XIC(FV_R2V2.CW.[CWD.FAULT]) XIC(Item_Faults_Are_Latched) ,XIC(FV_R2V2.CW.[CWD.HIGHLIGHT]) ] XIO(FV_R2V2.CW.[CWD.CHECKOFF]) XIO(Alarm_Reset) [OTE(FV_R2V2.CW.[CWD.FAULT]) ,ALMD(FV_R2V2_ALARM,0,0,0,0) ] ,XIC(FV_R2V2.CW.[CWD.OUTPUT]) OTE(FV_R2V2.CW.[CWD.PREVSCAN]) ,XIC(FV_R2V2.CW.[CWD.FAULT]) EQU(Scada_Valve_Fault_No,0) XIO(FV_R2V2.CW.[CWD.FAULTLOGGED]) [MOV(10001,Scada_Valve_Fault_No) ,OTL(FV_R2V2.CW.[CWD.FAULTLOGGED]) ] ];
   10: [NEQ(FV_AV5.DriveBits,0) OTE(FV_AV5.CW.[CWD.AUTODRV]) ,[XIC(FV_AV5.CW.[CWD.AUTODRV]) XIO(FV_AV5.CW.[CWD.MANUAL]) ,XIC(FV_AV5.CW.[CWD.MANDRV]) XIC(FV_AV5.CW.[CWD.MANUAL]) ] OTE(FV_AV5.CW.[CWD.OUTPUT]) ,XIC(FV_AV5.CW.[CWD.OUTPUT]) OTE(FV_AV5_DR) ,XIC(S:FS) [OTU(FV_AV1.CW.[CWD.MANUAL]) ,LEQ(FV_AV5.CheckTime,0) MOV(Default_Check_Time,FV_AV5.CheckTime) ] ,[[XIC(FV_AV5_O) XIO(Item_Simulation_Flag) ,XIC(Item_Simulation_Flag) XIC(FV_AV5.CW.[CWD.OUTPUT]) XIO(FV_AV5.CW.[CWD.SIMFAIL]) ] OTE(FV_AV5.CW.[CWD.OPENFB]) ,[XIC(FV_AV5_C) XIO(Item_Simulation_Flag) ,XIC(Item_Simulation_Flag) XIO(FV_AV5.CW.[CWD.OUTPUT]) XIO(FV_AV5.CW.[CWD.SIMFAIL]) ] OTE(FV_AV5.CW.[CWD.CLOSEDFB]) ] ,[XIC(FV_AV5.CW.[CWD.OUTPUT]) XIO(FV_AV5.CW.[CWD.PREVSCAN]) ,XIO(FV_AV5.CW.[CWD.OUTPUT]) XIC(FV_AV5.CW.[CWD.PREVSCAN]) ] CLR(FV_AV5.CheckTimer) ,XIC(One_Second_One_Scan) LES(FV_AV5.CheckTimer,FV_AV5.CheckTime) ADD(FV_AV5.CheckTimer,1,FV_AV5.CheckTimer) ,XIO(FV_AV5.CW.[CWD.FAULT]) OTU(FV_AV5.CW.[CWD.FAULTLOGGED]) ,[GEQ(FV_AV5.CheckTimer,FV_AV5.CheckTime) [XIC(FV_AV5.CW.[CWD.OUTPUT]) [XIO(FV_AV5.CW.[CWD.OPENFB]) ,XIC(FV_AV5.CW.[CWD.CLOSEDFB]) ] ,XIO(FV_AV5.CW.[CWD.OUTPUT]) [XIC(FV_AV5.CW.[CWD.OPENFB]) ,XIO(FV_AV5.CW.[CWD.CLOSEDFB]) ] ] ,XIC(FV_AV5.CW.[CWD.FAULT]) XIC(Item_Faults_Are_Latched) ,XIC(FV_AV5.CW.[CWD.HIGHLIGHT]) ] XIO(FV_AV5.CW.[CWD.CHECKOFF]) XIO(Alarm_Reset) [OTE(FV_AV5.CW.[CWD.FAULT]) ,ALMD(FV_AV5_ALARM,0,0,0,0) ] ,XIC(FV_AV5.CW.[CWD.OUTPUT]) OTE(FV_AV1.CW.[CWD.PREVSCAN]) ,XIC(FV_AV5.CW.[CWD.FAULT]) EQU(Scada_Valve_Fault_No,0) XIO(FV_AV5.CW.[CWD.FAULTLOGGED]) [MOV(10005,Scada_Valve_Fault_No) ,OTL(FV_AV5.CW.[CWD.FAULTLOGGED]) ] ];
   // Yeast Press AV2 (Blunger Pump Solenoid)
   11: [NEQ(YP_AV2.DriveBits,0) OTE(YP_AV2.CW.[CWD.AUTODRV]) ,[XIC(YP_AV2.CW.[CWD.AUTODRV]) XIO(YP_AV2.CW.[CWD.MANUAL]) ,XIC(YP_AV2.CW.[CWD.MANDRV]) XIC(YP_AV2.CW.[CWD.MANUAL]) ] OTE(YP_AV2.CW.[CWD.OUTPUT]) ,XIC(YP_AV2.CW.[CWD.OUTPUT]) OTE(YP_AV2_DR) ,XIC(S:FS) [OTU(YP_AV2.CW.[CWD.MANUAL]) ,LEQ(YP_AV2.CheckTime,0) MOV(Default_Check_Time,YP_AV2.CheckTime) ] ,[[XIC(YP_AV2_O) XIO(Item_Simulation_Flag) ,XIC(Item_Simulation_Flag) XIC(YP_AV2.CW.[CWD.OUTPUT]) XIO(YP_AV2.CW.[CWD.SIMFAIL]) ] OTE(YP_AV2.CW.[CWD.OPENFB]) ,[XIO(YP_AV2_O) XIO(Item_Simulation_Flag) ,XIC(Item_Simulation_Flag) XIO(YP_AV2.CW.[CWD.OUTPUT]) XIO(YP_AV2.CW.[CWD.SIMFAIL]) ] OTE(YP_AV2.CW.[CWD.CLOSEDFB]) ] ,[XIC(YP_AV2.CW.[CWD.OUTPUT]) XIO(YP_AV2.CW.[CWD.PREVSCAN]) ,XIO(YP_AV2.CW.[CWD.OUTPUT]) XIC(YP_AV2.CW.[CWD.PREVSCAN]) ] CLR(YP_AV2.CheckTimer) ,XIC(One_Second_One_Scan) LES(YP_AV2.CheckTimer,YP_AV2.CheckTime) ADD(YP_AV2.CheckTimer,1,YP_AV2.CheckTimer) ,XIO(YP_AV2.CW.[CWD.FAULT]) OTU(YP_AV2.CW.[CWD.FAULTLOGGED]) ,[GEQ(YP_AV2.CheckTimer,YP_AV2.CheckTime) [XIC(YP_AV2.CW.[CWD.OUTPUT]) [XIO(YP_AV2.CW.[CWD.OPENFB]) ,XIC(YP_AV2.CW.[CWD.CLOSEDFB]) ] ,XIO(YP_AV2.CW.[CWD.OUTPUT]) [XIC(YP_AV2.CW.[CWD.OPENFB]) ,XIO(YP_AV2.CW.[CWD.CLOSEDFB]) ] ] ,XIC(YP_AV2.CW.[CWD.FAULT]) XIC(Item_Faults_Are_Latched) ,XIC(YP_AV2.CW.[CWD.HIGHLIGHT]) ] XIO(YP_AV2.CW.[CWD.CHECKOFF]) XIO(Alarm_Reset) [OTE(YP_AV2.CW.[CWD.FAULT]) ,ALMD(YP_AV2_ALARM,0,0,0,0) ] ,XIC(YP_AV2.CW.[CWD.OUTPUT]) OTE(YP_AV2.CW.[CWD.PREVSCAN]) ];
END_ROUTINE
